// TIA Portal project "XSFW_TIA32801_A0" (V15.1)

(* hardware
DEVICE "Estación SIMATIC 1200_1"  S71200.Device
   slot 0: "Rack S7-1200"  Rack  V1.0
   slot 1: "PLC_1"  CPU 1214C DC/DC/DC  6ES7 214-1AG40-0XB0  V4.3
   slot 2: "DI16/DQ16 x 24V DC_1"  6ES7 223-1BL30-0XB0  V1.0
   slot 3: "DI 8x24VDC_1"  6ES7 221-1BF32-0XB0  V2.0
DEVICE "HMI_1"  KTP700 Basic PN
   slot 0: "HMI_1"  KTP700 Basic PN  6AV2 123-2GB03-0AX0  15.1.0.0
   slot 1: "HMI_RT_1"  KTP700 Basic PN  6AV2 123-2GB03-0AX0  15.1.0.0
   slot 5: "IE_CP_1"  PROFINET Interface  IE_CP  15.0.1.0
      slot 1: "PROFINET_Interfaz_1"  PROFINET Interface
         slot 1: "PORT_1"  Port  1.0.0.0
*)

// ===== PLC "PLC_1"  CPU 1214C DC/DC/DC =====

VAR_GLOBAL   // PLC tag table "Constantes del sistema"
   "Encoder" AT %ID1000 : DWord;   // Almacena el valor actual del encoder
   "System_Byte" AT %MB61 : Byte;
   "Clock_Byte" AT %MB60 : Byte;
   "Marca del sistema" AT %M61.0 : Bool;   // marca del sistema
   "Marca de ciclo" AT %M60.0 : Bool;   // Genera una luz titilante de 10 hz
   "No entrega caja" AT %M100.0 : Bool;
   "No libera salida" AT %M100.1 : Bool;
   "HMI_Hab. Falla caja trab." AT %M100.2 : Bool;
   "Tag_4" AT %M100.3 : Bool;
   "Tag_5" AT %M100.4 : Bool;
   "Tag_6" AT %M100.5 : Bool;
   "Tag_7" AT %M100.6 : Bool;
   "Tag_8" AT %M100.7 : Bool;
   "Tag_9" AT %M101.0 : Bool;
   "bit 1 de Reg_A" AT %M101.1 : Bool;
   "Tag_11" AT %M101.2 : Bool;
   "Tag_12" AT %M101.3 : Bool;
   "Tag_13" AT %M101.4 : Bool;
   "Tag_14" AT %M101.5 : Bool;
   "Tag_15" AT %M101.6 : Bool;
   "Tag_16" AT %M101.7 : Bool;
   "bit 0 de Reg_B" AT %M102.0 : Bool;
   "Tag_18" AT %M102.1 : Bool;
   "Tag_19" AT %M102.2 : Bool;
   "Tag_20" AT %M102.3 : Bool;
   "Tag_21" AT %M102.4 : Bool;
   "Tag_22" AT %M102.5 : Bool;
   "Tag_23" AT %M102.6 : Bool;
   "Tag_24" AT %M102.7 : Bool;
   "Tag_25" AT %M103.0 : Bool;
   "Tag_26" AT %M103.1 : Bool;
   "Tag_27" AT %M103.2 : Bool;
   "Tag_28" AT %QB0 : Byte;
   "UNO" AT %M27.0 : Bool;
   "CERO" AT %M27.1 : Bool;
   "Marca ciclo alim cartones" AT %M60.1 : Bool;   // es una marca de ciclo de 5 hz para manejar el alim de cartones
   "Tag_29" AT %M60.2 : Bool;
   "Tag_30" AT %M60.5 : Bool;
   "Tag_31" AT %MD300 : DWord;
   "Valor encoder pusher salida" AT %MD350 : DWord;
   "Tag_32" AT %E0.7 : Bool;
   "Tag_33" AT %M36.4 : Bool;
   "Reg_A" AT %MB101 : Byte;
   "Reg_B" AT %MB102 : Byte;
   "Tag_1" AT %I34.2 : Bool;
END_VAR

VAR_GLOBAL   // PLC tag table "Pusher"
   "iSNSpush_atras" AT %I33.2 : Bool;   // Detecta Pusher atrás
   "iSNSpush_adel" AT %I0.2 : Bool;   // Detecta Pusher adelante
   "iSNSalp" AT %I1.0 : Bool;   // Sensor área de recorrido libre del pusher
   "oM_pusher" AT %Q32.3 : Bool;   // Activa el pusher
   "oPusher_out" AT %Q33.5 : Bool;   // Activa válvula del Cilindro del pusher
END_VAR

VAR_GLOBAL   // PLC tag table "brazo de succion"
   "iSNS_bs_abajo" AT %I33.6 : Bool;   // Detecta cuando el brazo de succión está abajo
   "iSNS_bs_arriba" AT %I33.7 : Bool;   // Detecta cuando el brazo de succión está arriba
   "oM_brazo_succión" AT %Q32.2 : Bool;   // Activa el brazo de succión
   "oVálvula_Succión" AT %Q33.0 : Bool;   // Activa valvula chupetes succionadores
END_VAR

VAR_GLOBAL   // PLC tag table "Pinza"
   "oPinza" AT %Q33.6 : Bool;   // Activa válvula Brazos tipo pinza que cierran las solapas inferiores de la caja
END_VAR

VAR_GLOBAL   // PLC tag table "agarra solapa, cierra solapa, alimentador de caja,retenedores"
   "oAgarra_solapas" AT %Q33.1 : Bool;   // Activa válvula brazos agarra solapas
   "oCierra_solapa" AT %Q33.2 : Bool;   // Activa válvula brazo cierra solapa
   "oRetB" AT %Q33.3 : Bool;   // Activa válvula Retenedor de caja en sector B
   "oRetC" AT %Q33.7 : Bool;   // Activa válvula Retenedor de cajas en sector C
   "oAlim_cart" AT %Q0.0 : Bool;   // Válvula Alimentación automática de cartones
   "iSNS_nivel_bajo_cartones" AT %I33.0 : Bool;   // Detecta nivel bajo de cartones
END_VAR

VAR_GLOBAL   // PLC tag table "Encoladora"
   "iSNS_carton en area de colado" AT %I33.3 : Bool;   // Detecta el cartón en sector de colado
   "iK_encol_on" AT %I33.1 : Bool;   // Encoladora encendida y caliente (tarda 45 min en calentar)
   "iSNSpegamento en depósito" AT %I1.2 : Bool;   // Detecta pegamento en depósito
   "oBoquilla_Encoladora" AT %Q33.4 : Bool;   // Activa Boquilla encoladora
END_VAR

VAR_GLOBAL   // PLC tag table "Area de salida"
   "iSNScaja_trab" AT %I1.4 : Bool;   // Detecta cuando la caja cae a la cinta de salida
   "iSnsCajaCerrada" AT %I1.5 : Bool;   // Detecta si la caja no se abrio cuando bajo a la cadena
   "oM_cinta_sal" AT %Q32.4 : Bool;   // Activa la cinta de salida
   "iSNScaja_acum" AT %I0.4 : Bool;   // detecta cajas acumuladas
END_VAR

VAR_GLOBAL   // PLC tag table "Cinta y encoder"
   "iFaseA" AT %I0.0 : Bool;   // fase A del encoder
   "iFaseB" AT %I0.1 : Bool;   // fase B del encoder
   "iFase0" AT %I0.3 : Bool;   // fase 0 del encoder, detecta cuando se cumplió una vuelta
   "oM_cinta_principal" AT %Q32.0 : Bool;   // Activa el motor de la cinta principal
END_VAR

VAR_GLOBAL   // PLC tag table "auxiliares para almacenar flancos"
   "Guarda flanco subida caja acum" AT %M80.0 : Bool;   // almacena valor anterior del sensor caja acumulada
   "Guarda flanco bajada caja acum" AT %M80.1 : Bool;   // almacena valor anterior del sensor caja acumulada
   "Guarda flanco bajada caja trab" AT %M80.2 : Bool;   // almacena valor anterior del sensor caja trabada
   "Guarda flanco subida caja trab" AT %M80.3 : Bool;   // almacena valor anterior del sensor caja trabada
   "Guarda flanco brazo succión arriba" AT %M80.4 : Bool;   // Almacena el estado anterior del sensor
   "Guarda flanco subida area encolado" AT %M80.5 : Bool;
   "Guarda flanco bajada area encolado" AT %M80.6 : Bool;
   "Guarda flanco pulsador averia/reposicion" AT %M80.7 : Bool;
   "Guarda flanco subida pulsador marcha" AT %M81.0 : Bool;
   "Guarda flanco subida pulsador avería/reposición" AT %M81.1 : Bool;
   "Guarda flanco subida pulsador Parada" AT %M81.2 : Bool;
   "fls_Averiarep" AT %M81.3 : Bool;
   "fls_M" AT %M81.4 : Bool;
   "fls_Area_encol_sub" AT %M81.5 : Bool;
   "fls_Area_encol_baj" AT %M81.6 : Bool;
   "Guarda flanco Marcha desde panel" AT %M81.7 : Bool;
   "Guarda flanco modo manual" AT %M82.0 : Bool;
   "fls_Modomanual" AT %M82.1 : Bool;   // Pulsador desde panel para comenzar modo manual
   "Guarda flanco bajada alim cart" AT %M82.2 : Bool;
   "Guarda flanco de bajada sns brazo abajo" AT %M82.3 : Bool;
END_VAR

VAR_GLOBAL   // PLC tag table "Pulsadores y selectores"
   "iM" AT %I32.5 : Bool;   // Pulsador de Marcha
   "iP" AT %I32.6 : Bool;   // Pulsador de Parada
   "iS_automat" AT %I33.4 : Bool;   // Selector modo automático
   "iS_Probar" AT %I33.5 : Bool;   // Selector modo test
   "iS_cinta_salida_on" AT %I1.3 : Bool;   // Selectora on/off de la cinta de salida
END_VAR

VAR_GLOBAL   // PLC tag table "Seguridad"
   "iEmergencia" AT %I32.1 : Bool;   // Ventanas cerradas y emerg off
   "iAveria-reposicion" AT %I32.2 : Bool;   // Repone avería
   "iTermicas_mev" AT %I32.3 : Bool;   // Térmicas del motor, encoladora, bomba
   "iTermicas_pbs" AT %I32.4 : Bool;   // Térmicas del brazo de succión y pusher
   "iSNSproteccion_torque" AT %I0.5 : Bool;   // Sensor Protección de torque motor principal cinta
   "oLinea-emergencia" AT %Q32.7 : Bool;   // Salida a línea de emergencia
END_VAR

VAR_GLOBAL   // PLC tag table "voltage de control"
   "iEnable" AT %I32.0 : Bool;   // Voltage de control
END_VAR

VAR_GLOBAL   // PLC tag table "Otros"
   "k_EXT" AT %I1.1 : Bool;   // enable suction arm from EXT input
   "oQuick_out" AT %Q0.1 : Bool;   // ?
   "oSep_fing" AT %Q0.4 : Bool;   // ?
   "oPacker" AT %Q0.3 : Bool;   // En teoría se habilita luego que pulsa Marcha
   "desactivar" AT %M50.0 : Bool;
END_VAR

VAR_GLOBAL   // PLC tag table "Bomba de vacio"
   "oM_bomba" AT %Q32.1 : Bool;   // Activa la bomba de vacío
END_VAR

VAR_GLOBAL   // PLC tag table "Luces"
   "oLmpR" AT %Q32.5 : Bool;   // Lámpara para indicar parada y fallas de cualquier índole
   "oLmpV" AT %Q32.6 : Bool;   // Lámpara para indicar marcha
END_VAR

VAR_GLOBAL   // PLC tag table "Estados"
   "DS1" AT %MD0 : DWord;   // Variable tipo Word. Almacena los 12 Estados del proceso
   "1s1" AT %M0.0 : Bool;   // Estado 1: Reposo
   "1s2" AT %M0.1 : Bool;   // Estado 2: Activa Cinta ppal
   "1s3" AT %M0.2 : Bool;   // Estado 3: Activar retenedores de caja
   "1s4" AT %M0.3 : Bool;   // Estado 4: Desactivar Cinta ppal
   "1s5" AT %M0.4 : Bool;   // Estado 5: Activar Pusher y Pinza
   "1s6" AT %M0.5 : Bool;   // Estado 6: Activar Cilindro neumático Pusher
   "1s7" AT %M0.6 : Bool;   // Estado 7: Desactivar Pinza y Cilindro Pusher
   "1s8" AT %M0.7 : Bool;   // Estado 8: Área libre de Pusher
   "1s9" AT %M1.0 : Bool;   // Estado 9: Fin Etapa Pusher
   "1s10" AT %M1.1 : Bool;
   "1s11" AT %M1.2 : Bool;
   "1s12" AT %M1.3 : Bool;
   "DS2" AT %MD4 : DWord;
   "2s1" AT %M4.0 : Bool;   // Estado 8: Activar retenedores de caja
   "2s2" AT %M4.1 : Bool;   // Estado 9: Desactivar cinta
   "2s3" AT %M4.2 : Bool;   // Estado 10: Activa Pusher, Pinza y Cierra solapa
   "2s4" AT %M4.3 : Bool;   // Estado 11: Cilindro Pusher Afuera
   "2s5" AT %M4.4 : Bool;   // Estado 12: Desactivar Cilindro Pusher, Pinza y Cierra solapa
   "2s6" AT %M4.5 : Bool;   // Estado 13: Fin Pusher
   "2s7" AT %M4.6 : Bool;   // Estado 14: Area liberada del Pusher
   "2s8" AT %M4.7 : Bool;
   "2s9" AT %M5.0 : Bool;
   "2s10" AT %M5.1 : Bool;
   "2s11" AT %M5.2 : Bool;
   "2s12" AT %M5.3 : Bool;
   "2s13" AT %M5.4 : Bool;
   "2s14" AT %M5.5 : Bool;
   "2s15" AT %M5.6 : Bool;
   "2s16" AT %M5.7 : Bool;
   "2s17" AT %M6.0 : Bool;
   "2s18" AT %M6.1 : Bool;
   "2s19" AT %M6.2 : Bool;
   "2s20" AT %M6.3 : Bool;
   "2s21" AT %M6.4 : Bool;
   "2s22" AT %M6.5 : Bool;
   "2s23" AT %M6.6 : Bool;
   "2s24" AT %M6.7 : Bool;
   "2s25" AT %M7.0 : Bool;
   "2s26" AT %M7.1 : Bool;
   "2s27" AT %M7.2 : Bool;
   "2s28" AT %M7.3 : Bool;
   "2s29" AT %M7.4 : Bool;
   "2s30" AT %M7.5 : Bool;
   "2s31" AT %M7.6 : Bool;
   "2s32" AT %M7.7 : Bool;
   "1s13" AT %M1.4 : Bool;
   "1s14" AT %M1.5 : Bool;
   "1s15" AT %M1.6 : Bool;
   "1s16" AT %M1.7 : Bool;
   "1s17" AT %M2.0 : Bool;
   "1s18" AT %M2.1 : Bool;
   "1s19" AT %M2.2 : Bool;
   "1s20" AT %M2.3 : Bool;   // Estado de Alarmas
   "1s21" AT %M2.4 : Bool;   // Estado de parada
   "1s22" AT %M2.5 : Bool;   // Cajas acumuladas
   "1s23" AT %M2.6 : Bool;
   "1s24" AT %M2.7 : Bool;
   "1s25" AT %M3.0 : Bool;
   "1s26" AT %M3.1 : Bool;
   "1s27" AT %M3.2 : Bool;
   "1s28" AT %M3.3 : Bool;
   "1s29" AT %M3.4 : Bool;
   "1s30" AT %M3.5 : Bool;
   "1s31" AT %M3.6 : Bool;
   "1s32" AT %M3.7 : Bool;
END_VAR

VAR_GLOBAL   // PLC tag table "Concatenadores"
   "DC1" AT %MD8 : DWord;
   "1c1" AT %M8.0 : Bool;   // Ir a Estado 1: Reposo
   "1c2" AT %M8.1 : Bool;   // Ir a estado 2: Activa Cinta ppal
   "1c3" AT %M8.2 : Bool;   // Ir a estado 3: Activar retenedores de caja
   "1c4" AT %M8.3 : Bool;   // Ir estado 4: Desactivar Cinta ppal
   "1c5" AT %M8.4 : Bool;   // Ir a estado 5: Activar Pusher y Pinza
   "1c6" AT %M8.5 : Bool;   // Ir a estado 6: Activar cilindro neumático Pusher
   "1c7" AT %M8.6 : Bool;   // Ir a estado 7: Desactivar Pinza y Cilindro Pusher
   "DC2" AT %MD12 : DWord;
   "2c1" AT %M12.0 : Bool;   // Ir a Estado 8: Activar retenedores de caja
   "2c2" AT %M12.1 : Bool;   // Ir a Estado 9: Desactivar cinta
   "2c3" AT %M12.2 : Bool;   // Ir a Estado 10: Activa Pusher, Pinza y Cierra solapa
   "2c4" AT %M12.3 : Bool;   // Ir a Estado 11: Cilindro Pusher afuera
   "2c5" AT %M12.4 : Bool;   // Ir a Estado 12: Desactivar Cilindro Pusher, Pinza y Cierra solapa
   "2c6" AT %M12.5 : Bool;   // Ir a Estado 13: Fin Pusher
   "2c7" AT %M12.6 : Bool;   // Ir a Estado 14: Area liberada del Pusher
   "1c8" AT %M8.7 : Bool;   // Ir a Estado 8: Área libre de Pusher
   "1c9" AT %M9.0 : Bool;   // Ir a Estado 9: Fin etapa Pusher
   "1c10" AT %M9.1 : Bool;
   "1c11" AT %M9.2 : Bool;
   "1c12" AT %M9.3 : Bool;
   "1c13" AT %M9.4 : Bool;
   "1c14" AT %M9.5 : Bool;
   "1c15" AT %M9.6 : Bool;
   "1c16" AT %M9.7 : Bool;
   "1c17" AT %M10.0 : Bool;
   "1c18" AT %M10.1 : Bool;
   "1c19" AT %M10.2 : Bool;
   "1c20" AT %M10.3 : Bool;
   "1c21" AT %M10.4 : Bool;
   "1c22" AT %M10.5 : Bool;
   "1c23" AT %M10.6 : Bool;
   "1c24" AT %M10.7 : Bool;
   "1c25" AT %M11.0 : Bool;
   "1c26" AT %M11.1 : Bool;
   "1c27" AT %M11.2 : Bool;
   "1c28" AT %M11.3 : Bool;
   "1c29" AT %M11.4 : Bool;
   "1c30" AT %M11.5 : Bool;
   "1c31" AT %M11.6 : Bool;
   "1c32" AT %M11.7 : Bool;
   "2c8" AT %M12.7 : Bool;
   "2c9" AT %M13.0 : Bool;
   "2c10" AT %M13.1 : Bool;
   "2c11" AT %M13.2 : Bool;
   "2c12" AT %M13.3 : Bool;
   "2c13" AT %M13.4 : Bool;
   "2c14" AT %M13.5 : Bool;
   "2c15" AT %M13.6 : Bool;
   "2c16" AT %M13.7 : Bool;
   "2c17" AT %M14.0 : Bool;
   "2c18" AT %M14.1 : Bool;
   "2c19" AT %M14.2 : Bool;
   "2c20" AT %M14.3 : Bool;
   "2c21" AT %M14.4 : Bool;
   "2c22" AT %M14.5 : Bool;
   "2c23" AT %M14.6 : Bool;
   "2c24" AT %M14.7 : Bool;
   "2c25" AT %M15.0 : Bool;
   "2c26" AT %M15.1 : Bool;
   "2c27" AT %M15.2 : Bool;
   "2c28" AT %M15.3 : Bool;
   "2c29" AT %M15.4 : Bool;
   "2c30" AT %M15.5 : Bool;
   "2c31" AT %M15.6 : Bool;
   "2c32" AT %M15.7 : Bool;
END_VAR

VAR_GLOBAL   // PLC tag table "Marcas"
   "Marcha" AT %M20.0 : Bool;   // marca "Iniciar proceso"
   "Activar desplazador" AT %M20.1 : Bool;   // marca "activar cilindro alimentador"
   "Activa_cinta_salida" AT %M20.2 : Bool;   // marca " activa cinta de salida"
   "HMI_Hab_Falla_Caja_Caida" AT %M20.3 : Bool;   // Cajas acumuladas en la cinta de salida
   "Interrumpir" AT %M20.4 : Bool;   // Interrumpe el proceso
   "Activa pinza" AT %M20.5 : Bool;   // Activa la pinza
   "Activa cierra solapa" AT %M20.6 : Bool;   // Activa el cierra solapa
   "Activa bomba" AT %M20.7 : Bool;   // Activa la bomba de vacío
   "Activa brazo_succion" AT %M21.0 : Bool;   // Activa el motor del brazo de succión
   "Pusher-atras-ok" AT %M21.2 : Bool;   // Confirma que el pusher tocó el sensor de atrás
   "Pusher-adelante-ok" AT %M21.3 : Bool;   // Confirma que el pusher tocó el sensor adelante
   "Area libre del pusher" AT %M21.4 : Bool;   // Confirma que se activó el sensor
   "Ya buscó caja" AT %M21.5 : Bool;   // Confirma que el brazo tomó una caja
   "Activa succionadores" AT %M21.6 : Bool;   // Marca que activa los chupetes succionadores
   "No salió caja" AT %M21.7 : Bool;   // Indica que la caja no salió del rango del brazo de succión
   "Aux1" AT %M22.0 : Bool;   // auxiliar para los registros SR
   "Aux2" AT %M22.1 : Bool;   // auxiliar para los registros SR
   "Aux3" AT %M22.2 : Bool;   // auxiliar para los registros SR
   "Aux4" AT %M22.3 : Bool;   // auxiliar para los registros SR
   "Aux5" AT %M22.4 : Bool;   // auxiliar para los registros SR
   "Encolado fallido o falla en sensor" AT %M23.0 : Bool;   // Indica que el encolado se realizó correctamente, se da cuuando NO se da falla en encolado
   "Rearmar" AT %M23.1 : Bool;   // Se activa cuando se presiona el pulsador de avería/reposición
   "Falla en pusher" AT %M23.2 : Bool;   // Indica que hubo una falla en el pusher
   "Alarmas pusher" AT %M23.3 : Bool;   // Agrupa las alarmas del pusher
   "Alarmas brazo de succión" AT %M23.4 : Bool;   // Agrupa las alarmas del brazo de succión
   "Alarmas emergencia y térmicas" AT %M23.5 : Bool;   // Agrupa las alarmas de la serie térmicas y serie emergencia y ventanas
   "Alarmas cinta" AT %M23.6 : Bool;   // Agrupa las alarmas de la cinta
   "Alarmas salida y alim de cartones" AT %M23.7 : Bool;   // Agrupa las alarmas de la salida de la máquina (caja trabada) y alimentación de cartones
   "Cajas acumuladas en salida" AT %M24.0 : Bool;   // Detecta acumulación de cajas en la cinta salida interrumpiendo el proceso
   "Aux6" AT %M24.1 : Bool;
   "Alarmas encoladora" AT %M24.2 : Bool;
   "Serie de Alarmas" AT %M24.3 : Bool;
   "Habilita modo Probar" AT %M24.4 : Bool;
   "Tiempo de encolado solapa 1" AT %M24.5 : Bool;
   "Tiempo de encolado solapa2" AT %M24.6 : Bool;
   "Serie de fallas" AT %M24.7 : Bool;
   "Rearme desde panel" AT %M25.0 : Bool;
   "Emergencia desde panel" AT %M25.1 : Bool;
   "Valor del encoder" AT %MD180 : DWord;
   "Parada" AT %M25.2 : Bool;
   "Marcha desde panel" AT %M25.3 : Bool;
   "Modo Manual" AT %M25.4 : Bool;   // Cuando no está en modo probar ni en modo aut, está en modo manual
   "Resetear cajas armadas" AT %M25.5 : Bool;
   "Valor cantidad de cajas armadas" AT %MD120 : DWord;
   "Valor de referencia cajas armadas" AT %M25.6 : Bool;
   "Aux7" AT %M25.7 : Bool;
   "Solapa en área de encolado" AT %M26.0 : Bool;
   "Solapa fuera del area de encolado" AT %M26.1 : Bool;
   "Valorexp de contaje para calcular encolado x" AT %MD150 : DWord;
   "Exp Almacena el valor encolado experimental" AT %MD170 : DWord;
   "Exp marca de prueba fase 0" AT %M26.2 : Bool;   // Esta marca sólo me sirve a mi para ver si la fase 0 efectiv se activa
   "Impedir falla" AT %M26.3 : Bool;
   "Boton activar fingers" AT %M26.4 : Bool;
   "Botón packer" AT %M26.5 : Bool;
   "Boton quick out" AT %M26.6 : Bool;
   "Exp valor del encoder para calc encolado" AT %MD220 : DWord;
   "Exp marca aux id118" AT %M22.5 : Bool;
   "Pulsador modo manual" AT %M22.6 : Bool;   // Cada vez que se pulsa, se lleva a cabo un ciclo de la armadora
   "Aviso de cinta descalibrada probar" AT %M22.7 : Bool;
   "Habilitar brazo manual" AT %M26.7 : Bool;
   "Aux alim cart" AT %M27.2 : Bool;
   "Aux alim cart 2" AT %M27.3 : Bool;
   "Iniciar temp alim cart" AT %M27.4 : Bool;
   "Recuerda paso pusher" AT %M27.5 : Bool;
   "Auxiliar encoder exp" AT %M27.6 : Bool;
   "Aux9" AT %M27.7 : Bool;
   "Punto neutro" AT %M28.0 : Bool;
   "Aux10" AT %M28.1 : Bool;
   "Aux11" AT %M28.2 : Bool;
   "Delay cierra solapa" AT %M28.3 : Bool;
   "Delay brazo" AT %M28.4 : Bool;
   "Delay brazo 2" AT %M28.5 : Bool;
   "Aux12" AT %M28.6 : Bool;
   "Auxencol1" AT %M28.7 : Bool;
   "Auxencol2" AT %M29.0 : Bool;
   "Guarda flanco bajada averi rep delay" AT %M29.1 : Bool;
   "Rearme delay" AT %M29.2 : Bool;
   "Delaymarcha" AT %M29.3 : Bool;
   "Guarda flanco delay  marcha" AT %M29.4 : Bool;
   "Parar proceso" AT %M29.5 : Bool;
   "Espera caja" AT %M29.6 : Bool;
   "Guarda flanco punto m" AT %M29.7 : Bool;
   "Parar brazo" AT %M34.0 : Bool;
   "Flanco 2" AT %M34.1 : Bool;
   "Esperar cinta" AT %M34.2 : Bool;
   "Flanco p atras" AT %M34.3 : Bool;
   "Flanco nivel bajo" AT %M34.4 : Bool;
   "Retrasa nivel bajo c" AT %M34.5 : Bool;
   "Fls sns b abajo" AT %M34.6 : Bool;
   "Fls_bajada snsalp" AT %M34.7 : Bool;
   "Aux marca pusher" AT %M35.0 : Bool;
   "Aux acaja acum" AT %M35.1 : Bool;
   "Aux17" AT %M35.2 : Bool;
   "Aux caja trab" AT %M35.3 : Bool;
   "Marca aux" AT %M35.4 : Bool;
   "Fsnsalp" AT %M35.5 : Bool;
   "Xsnsalp" AT %M35.6 : Bool;
   "FallaSnsAtras" AT %M35.7 : Bool;
   "F1s8" AT %M36.0 : Bool;
   "X1s8" AT %M36.1 : Bool;
   "Flanco_PusherAtras" AT %M36.2 : Bool;
   "FlancoAtras_Detectado" AT %M36.3 : Bool;
END_VAR

VAR_GLOBAL   // PLC tag table "Prioritarias"
   "1p1" AT %M16.0 : Bool;
   "DP1" AT %MD16 : DWord;
   "1p2" AT %M16.1 : Bool;
   "1p3" AT %M16.2 : Bool;
   "1p4" AT %M16.3 : Bool;
   "DP2" AT %MD30 : DWord;
   "2p1" AT %M30.0 : Bool;
   "2p2" AT %M30.1 : Bool;
   "2p3" AT %M30.2 : Bool;
   "2p4" AT %M30.3 : Bool;
   "2p5" AT %M30.4 : Bool;
   "2p6" AT %M30.5 : Bool;
   "1p8" AT %M16.7 : Bool;
   "1p9" AT %M17.0 : Bool;
   "1p5" AT %M16.4 : Bool;
   "1p6" AT %M16.5 : Bool;
   "1p7" AT %M16.6 : Bool;
   "1p10" AT %M17.1 : Bool;
   "1p11" AT %M17.2 : Bool;
   "1p12" AT %M17.3 : Bool;
   "1p13" AT %M17.4 : Bool;
   "1p14" AT %M17.5 : Bool;
   "1p15" AT %M17.6 : Bool;
   "1p16" AT %M17.7 : Bool;
   "1p17" AT %M18.0 : Bool;
   "1p18" AT %M18.1 : Bool;
   "1p19" AT %M18.2 : Bool;
   "1p20" AT %M18.3 : Bool;   // Prioritaria que para el proceso y necesita rearme
   "1p21" AT %M18.4 : Bool;   // Prioritaria que para el proceso y no necesita rearme
   "1p22" AT %M18.5 : Bool;   // Cajas acumuladas
   "1p23" AT %M18.6 : Bool;
   "1p24" AT %M18.7 : Bool;
   "1p25" AT %M19.0 : Bool;
   "1p26" AT %M19.1 : Bool;
   "1p27" AT %M19.2 : Bool;
   "1p28" AT %M19.3 : Bool;
   "1p29" AT %M19.4 : Bool;
   "1p30" AT %M19.5 : Bool;
   "1p31" AT %M19.6 : Bool;
   "1p32" AT %M19.7 : Bool;
END_VAR

VAR_GLOBAL   // PLC tag table "Modo probar"
   "MPbrazo de succión arriba" AT %M40.0 : Bool;   // levanta el brazo de succión
   "MPbrazo de succión abajo" AT %M40.1 : Bool;
   "MPlevanta brazo" AT %M40.2 : Bool;
   "MPbaja brazo" AT %M40.3 : Bool;
   "MPbotón Activa succión" AT %M40.4 : Bool;
   "MPsucciona caja" AT %M40.6 : Bool;
   "MPboton Activar bomba de vacío" AT %M40.7 : Bool;
   "MPbotón Activar encoladora" AT %M41.0 : Bool;
   "MPtiempo de encolado" AT %M41.1 : Bool;   // Encola por 2 segundos, independientemente si sigo presionando el botón
   "MPbotón alimentador de cartones" AT %M41.2 : Bool;
   "MPbotón Agarra solapas" AT %M41.3 : Bool;
   "MPbotón Cierra solapa" AT %M41.4 : Bool;
   "MPbotón Avanzar cinta" AT %M41.5 : Bool;
   "MPvalor actual del encoder" AT %MD200 : DWord;
   "MPbotón Avanzar cinta por tramos" AT %M41.6 : Bool;
   "MPActivar cinta" AT %M41.7 : Bool;
   "MPbotón activar pusher" AT %M42.0 : Bool;
   "MPActivar pusher" AT %M42.1 : Bool;
   "MPActivar cilindro pusher" AT %M42.2 : Bool;
   "MPguarda flanco subida ALP" AT %M42.3 : Bool;
   "MPActivar pinza" AT %M42.4 : Bool;
   "MPActiva bomba de vacío" AT %M42.5 : Bool;
   "MPActiva encola" AT %M42.6 : Bool;
   "MPActiva alimentación cartones" AT %M42.7 : Bool;
   "MPActiva los agarra solapas" AT %M43.0 : Bool;
   "MPActiva el cierra solapa" AT %M43.1 : Bool;
   "MPActiva la cinta de salida de cajas" AT %M43.2 : Bool;
   "ModoProbar" AT %M43.3 : Bool;
   "MPbotón activar retenedores de caja" AT %M43.4 : Bool;
   "MPActiva retenedores de caja" AT %M43.5 : Bool;
   "MPAcomodar brazo de succión" AT %M43.6 : Bool;
   "MPReset cuenta modo probar" AT %M43.7 : Bool;
   "MPboton cilindro push" AT %M44.0 : Bool;
   "MPactivar cilindro push" AT %M44.1 : Bool;
END_VAR

DATA_BLOCK "Fallas"   // DB1
{ S7_Optimized_Access := 'FALSE' }
VERSION : 0.1
   VAR
      termicas1 : Bool;   // Térmicas de la bomba de vacío, motor ppal, encoladora.
      termicas2 : Bool;   // Térmicas brazo de succión y pusher.
      emergencia : Bool;   // Ventanas abiertas o pulsador de emergencia activado.
      "proteccion de torque" : Bool;   // Protección de torque motor ppal (atasco).
      "Falla en rele cadena" : Bool;   // Falla en sensor de caja en área de encolado.
      "Falla en sensores del Pusher" : Bool;   // Falla en sensor del pusher atrás
      "Sensor pusher hacia adelante" : Bool;   // Falla en sensor del pusher adelante
      falla_sns_bsucc_ar : Bool;   // Falla en sensor del brazo de succión arriba
      falla_sns_bsucc_ab : Bool;   // Falla en sensor del brazo de succión abajo
      "area de recorrido libre del pusher" : Bool;   // Falla en sensor del pusher área libre.
      falla_alim_cartones : Bool;   // Falla en sensor alimentador de cartones.
      falla_encoder : Bool;   // Falla en encoder
      "caja trabada a la salida" : Bool;   // Falla en sensor de caja trabada a la salida.
      "Incrongruencia pusher" : Bool;   // Incongruencia en sensores del pusher
      "Falla de programación prioritarias 1" : Bool;
      "Falla de programación concatenadoras 1" : Bool;
      "Falla de programación prioritarias 2" : Bool;
      "Falla de programación concatenadoras 2" : Bool;
      "Falla en sensor de encolado" : Bool;   // Falla en sensor área de encolado
      "Sin pegamento en el depósito" : Bool;   // Sin pegamento en el depósito
      "falla rele cadena" : Bool;
      "Falla de caja cerrada en cadena" : Bool;   // se activa si cae mal la caja
      "Reserva 1_2_1" : Bool;
      "Reserva 1_3_1" : Bool;
      "Reserva 1_4_1" : Bool;
      "Reserva 1_4_1_1" : Bool;
      "Reserva 1_4_1_2" : Bool;
      "Reserva 1_4_1_3" : Bool;
      "Reserva 1_4_1_4" : Bool;
      "Reserva 1_4_1_4_1" : Bool;
      "Reserva 1_4_1_4_1_1" : Bool;
      "Reserva 1_4_1_4_1_2" : Bool;
   END_VAR
BEGIN
END_DATA_BLOCK

DATA_BLOCK "HSC"   // DB4
{ S7_Optimized_Access := 'FALSE' }
VERSION : 0.1
   VAR
      "punto muerto" : Bool;   // Indica que la cinta está completamente detenida
      id118 : Bool;   // Cuando el encoder llega a contar 118 pulsos, apaga el motor
      "Se cumplio una vuelta" : Bool;   // Indica que el motor dió una vuelta completa
   END_VAR
BEGIN
END_DATA_BLOCK

DATA_BLOCK "datos de encolado"   // DB11
{ S7_Optimized_Access := 'FALSE' }
VERSION : 0.1
   VAR
      Iniciosol1cj1000 : DInt;
      finsol1cj1000 : DInt;
      Iniciosol2cj1000 : DInt;
      finsol2cj1000 : DInt;
      Iniciosol1cj1500 : DInt;
      finsol1cj1500 : DInt;
      Iniciosol2cj1500 : DInt;
      finsol2cj1500 : DInt;
      "selcaja1000/1500" : Bool;
   END_VAR
BEGIN
END_DATA_BLOCK

DATA_BLOCK "AjusteEncoder"   // DB17
{ S7_Optimized_Access := 'TRUE' }
VERSION : 0.1
   VAR
      Hab_Pusher : DInt := -10;   // 0
      Dhab_Pusher : DInt := 21;   // 21
      Reset_Val : DInt;
      Reset : Bool;
   END_VAR
BEGIN
END_DATA_BLOCK

DATA_BLOCK "Alarmas"   // DB19
{ S7_Optimized_Access := 'FALSE' }
VERSION : 0.1
   VAR
      termicas1 : Bool;   // Térmicas de la bomba de vacío, motor ppal, encoladora.
      termicas2 : Bool;   // Térmicas brazo de succión y pusher.
      emergencia : Bool;   // Ventanas abiertas o pulsador de emergencia activado.
      "proteccion de torque" : Bool;   // Protección de torque motor ppal (atasco).
      "falla en rele de cadena" : Bool;   // Falla en sensor de caja en área de encolado.
      "Falla en sensor atras del pusher" : Bool;   // Falla en sensor del pusher atrás
      "Sensor pusher hacia adelante" : Bool;   // Falla en sensor del pusher adelante
      falla_sns_bsucc_ar : Bool;   // Falla en sensor del brazo de succión arriba
      falla_sns_bsucc_ab : Bool;   // Falla en sensor del brazo de succión abajo
      "area de recorrido libre del pusher" : Bool;   // Falla en sensor del pusher área libre.
      falla_alim_cartones : Bool;   // Falla en sensor alimentador de cartones.
      falla_encoder : Bool;   // Falla en encoder
      "caja trabada a la salida" : Bool;   // Falla en sensor de caja trabada a la salida.
      "Incrongruencia pusher" : Bool;   // Incongruencia en sensores del pusher
      "Falla de programación prioritarias" : Bool;
      "Falla de programación concatenadoras" : Bool;
      "Falla de programación prioritarias 2" : Bool;
      "Falla de programación concatenadoras 2" : Bool;
      "Falla en sensor de encolado" : Bool;   // Falla en sensor área de encolado
      "Sin pegamento en el depósito" : Bool;   // Sin pegamento en el depósito
      "falla rele cadena" : Bool;
      "caja cerrada en cadena" : Bool;
      Reserva_9 : Bool;
      Reserva_10 : Bool;
      Reserva_11 : Bool;
      Reserva_12 : Bool;
      Reserva_13 : Bool;
      Reserva_14 : Bool;
      Reserva_15 : Bool;
      Reserva_15_1 : Bool;
      Reserva_15_1_1 : Bool;
      Reserva_15_1_2 : Bool;
   END_VAR
BEGIN
END_DATA_BLOCK

DATA_BLOCK "Tiempos"   // DB23
{ S7_Optimized_Access := 'FALSE' }
VERSION : 0.1
   VAR
      "Tiempo cierra sol" : DInt;
      "Tiempo espera brazo" : DInt;
      "tiempo cajas acum" : DInt;
      "Tiempo caja trabada" : DInt;
   END_VAR
BEGIN
END_DATA_BLOCK

// folder: System blocks/Program resources

DATA_BLOCK "Timer_DB2"   // DB2
{ S7_Optimized_Access := 'TRUE' }
AUTHOR : Simatic
FAMILY : IEC
NAME : IEC_TMR
VERSION : 1.0
// stored: InstanceOfName IEC_TIMER
"IEC_TIMER"
BEGIN
END_DATA_BLOCK

DATA_BLOCK "Timer_DB3"   // DB3
{ S7_Optimized_Access := 'TRUE' }
AUTHOR : Simatic
FAMILY : IEC
NAME : IEC_TMR
VERSION : 1.0
// stored: InstanceOfName IEC_TIMER
"IEC_TIMER"
BEGIN
END_DATA_BLOCK

DATA_BLOCK "Timer_DB5"   // DB5
{ S7_Optimized_Access := 'TRUE' }
AUTHOR : Simatic
FAMILY : IEC
NAME : IEC_TMR
VERSION : 1.0
// stored: InstanceOfName IEC_TIMER
"IEC_TIMER"
BEGIN
END_DATA_BLOCK

DATA_BLOCK "Timer_DB6"   // DB6
{ S7_Optimized_Access := 'TRUE' }
AUTHOR : Simatic
FAMILY : IEC
NAME : IEC_TMR
VERSION : 1.0
// stored: InstanceOfName IEC_TIMER
"IEC_TIMER"
BEGIN
END_DATA_BLOCK

DATA_BLOCK "Timer_DB7"   // DB7
{ S7_Optimized_Access := 'TRUE' }
AUTHOR : Simatic
FAMILY : IEC
NAME : IEC_TMR
VERSION : 1.0
// stored: InstanceOfName IEC_TIMER
"IEC_TIMER"
BEGIN
END_DATA_BLOCK

DATA_BLOCK "Timer_DB8"   // DB8
{ S7_Optimized_Access := 'TRUE' }
AUTHOR : Simatic
FAMILY : IEC
NAME : IEC_TMR
VERSION : 1.0
// stored: InstanceOfName IEC_TIMER
"IEC_TIMER"
BEGIN
END_DATA_BLOCK

DATA_BLOCK "Timer_DB9"   // DB9
{ S7_Optimized_Access := 'TRUE' }
AUTHOR : Simatic
FAMILY : IEC
NAME : IEC_TMR
VERSION : 1.0
// stored: InstanceOfName IEC_TIMER
"IEC_TIMER"
BEGIN
END_DATA_BLOCK

DATA_BLOCK "IEC_Timer_0_DB"   // DB10
{ S7_Optimized_Access := 'TRUE' }
AUTHOR : Simatic
FAMILY : IEC
NAME : IEC_TMR
VERSION : 1.0
// stored: InstanceOfName IEC_TIMER
"IEC_TIMER"
BEGIN
END_DATA_BLOCK

DATA_BLOCK "Timer_DB12"   // DB12
{ S7_Optimized_Access := 'TRUE' }
AUTHOR : Simatic
FAMILY : IEC
NAME : IEC_TMR
VERSION : 1.0
// stored: InstanceOfName IEC_TIMER
"IEC_TIMER"
BEGIN
END_DATA_BLOCK

DATA_BLOCK "Timer_DB13"   // DB13
{ S7_Optimized_Access := 'TRUE' }
AUTHOR : Simatic
FAMILY : IEC
NAME : IEC_TMR
VERSION : 1.0
// stored: InstanceOfName IEC_TIMER
"IEC_TIMER"
BEGIN
END_DATA_BLOCK

DATA_BLOCK "Timer_DB14"   // DB14
{ S7_Optimized_Access := 'TRUE' }
AUTHOR : Simatic
FAMILY : IEC
NAME : IEC_TMR
VERSION : 1.0
// stored: InstanceOfName IEC_TIMER
"IEC_TIMER"
BEGIN
END_DATA_BLOCK

DATA_BLOCK "Timer_DB15"   // DB15
{ S7_Optimized_Access := 'TRUE' }
AUTHOR : Simatic
FAMILY : IEC
NAME : IEC_TMR
VERSION : 1.0
// stored: InstanceOfName IEC_TIMER
"IEC_TIMER"
BEGIN
END_DATA_BLOCK

DATA_BLOCK "Contador_0"   // DB16
{ S7_Optimized_Access := 'TRUE' }
AUTHOR : SIMATIC
FAMILY : IEC
NAME : DCNTR
VERSION : 1.2
// stored: InstanceOfName IEC_DCOUNTER
"IEC_DCOUNTER"
BEGIN
END_DATA_BLOCK

DATA_BLOCK "Timer_DB18"   // DB18
{ S7_Optimized_Access := 'TRUE' }
AUTHOR : Simatic
FAMILY : IEC
NAME : IEC_TMR
VERSION : 1.0
// stored: InstanceOfName IEC_TIMER
"IEC_TIMER"
BEGIN
END_DATA_BLOCK

DATA_BLOCK "Timer_DB20"   // DB20
{ S7_Optimized_Access := 'TRUE' }
AUTHOR : Simatic
FAMILY : IEC
NAME : IEC_TMR
VERSION : 1.0
// stored: InstanceOfName IEC_TIMER
"IEC_TIMER"
BEGIN
END_DATA_BLOCK

DATA_BLOCK "Timer_DB21"   // DB21
{ S7_Optimized_Access := 'TRUE' }
AUTHOR : Simatic
FAMILY : IEC
NAME : IEC_TMR
VERSION : 1.0
// stored: InstanceOfName IEC_TIMER
"IEC_TIMER"
BEGIN
END_DATA_BLOCK

DATA_BLOCK "Timer_DB22"   // DB22
{ S7_Optimized_Access := 'TRUE' }
AUTHOR : Simatic
FAMILY : IEC
NAME : IEC_TMR
VERSION : 1.0
// stored: InstanceOfName IEC_TIMER
"IEC_TIMER"
BEGIN
END_DATA_BLOCK

DATA_BLOCK "Timer_DB24"   // DB24
{ S7_Optimized_Access := 'TRUE' }
AUTHOR : Simatic
FAMILY : IEC
NAME : IEC_TMR
VERSION : 1.0
// stored: InstanceOfName IEC_TIMER
"IEC_TIMER"
BEGIN
END_DATA_BLOCK

DATA_BLOCK "TOFF"   // DB26
{ S7_Optimized_Access := 'TRUE' }
AUTHOR : Simatic
FAMILY : IEC
NAME : IEC_TMR
VERSION : 1.0
// stored: InstanceOfName IEC_TIMER
"IEC_TIMER"
BEGIN
END_DATA_BLOCK

DATA_BLOCK "Desactivar Pusher"   // DB27
{ S7_Optimized_Access := 'TRUE' }
AUTHOR : Simatic
FAMILY : IEC
NAME : IEC_TMR
VERSION : 1.0
// stored: InstanceOfName IEC_TIMER
"IEC_TIMER"
BEGIN
END_DATA_BLOCK

DATA_BLOCK "Timer_DB30"   // DB30
{ S7_Optimized_Access := 'TRUE' }
AUTHOR : Simatic
FAMILY : IEC
NAME : IEC_TMR
VERSION : 1.0
// stored: InstanceOfName IEC_TIMER
"IEC_TIMER"
BEGIN
END_DATA_BLOCK

DATA_BLOCK "Timer_DB31"   // DB31
{ S7_Optimized_Access := 'TRUE' }
AUTHOR : Simatic
FAMILY : IEC
NAME : IEC_TMR
VERSION : 1.0
// stored: InstanceOfName IEC_TIMER
"IEC_TIMER"
BEGIN
END_DATA_BLOCK

// folder: (top level)

FUNCTION "Alimentador de cartones y cinta de salida" : Void   // FC1, LAD
TITLE = Desplaza una cinta que traslada los cartones hasta el brazo succionador.
{ S7_Optimized_Access := 'FALSE' }
VERSION : 0.1
BEGIN

REGION Network 1: Activa la cinta de salida
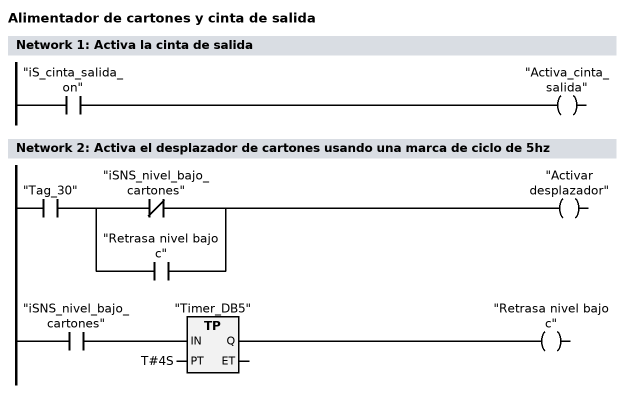
   RUNG wire#powerrail
      Contact( "iS_cinta_salida_on" )
      Coil( "Activa_cinta_salida" )
   END_RUNG
   // the same network as SCL:
   "Activa_cinta_salida" := "iS_cinta_salida_on";
END_REGION

REGION Network 2: Activa el desplazador de cartones usando una marca de ciclo de 5hz
   "Activar desplazador" := "Tag_30" AND (NOT "iSNS_nivel_bajo_cartones" OR "Retrasa nivel bajo c");
   "Timer_DB5".TP(IN := "iSNS_nivel_bajo_cartones", PT := T#4S);
   "Retrasa nivel bajo c" := "Timer_DB5".Q;
END_REGION
END_FUNCTION

FUNCTION "Tratamiento de Alarmas" : Void   // FC3, LAD
{ S7_Optimized_Access := 'TRUE' }
VERSION : 0.1
// Cada vez que ocurre una falla, cualquiera que fuese, se copia el estado de los bits de la doble palabra de "Fallas" a la doble palabra "Alarmas". Una vez resuelta la falla, se debe presionar "avería/reposición", lo cual generará un " reconocimiento de falla, que dará de baja la Alarma. A partir del segmento 4, agrupo las alarmas por función. Un grupo de alarmas para el pusher, uno para brazo de succión ,etc.
   VAR_TEMP
      "Alarmas presentes" : Word;
      Reconocimiento : Word;
   END_VAR
BEGIN

REGION Network 1: Reconocimiento/Reposición
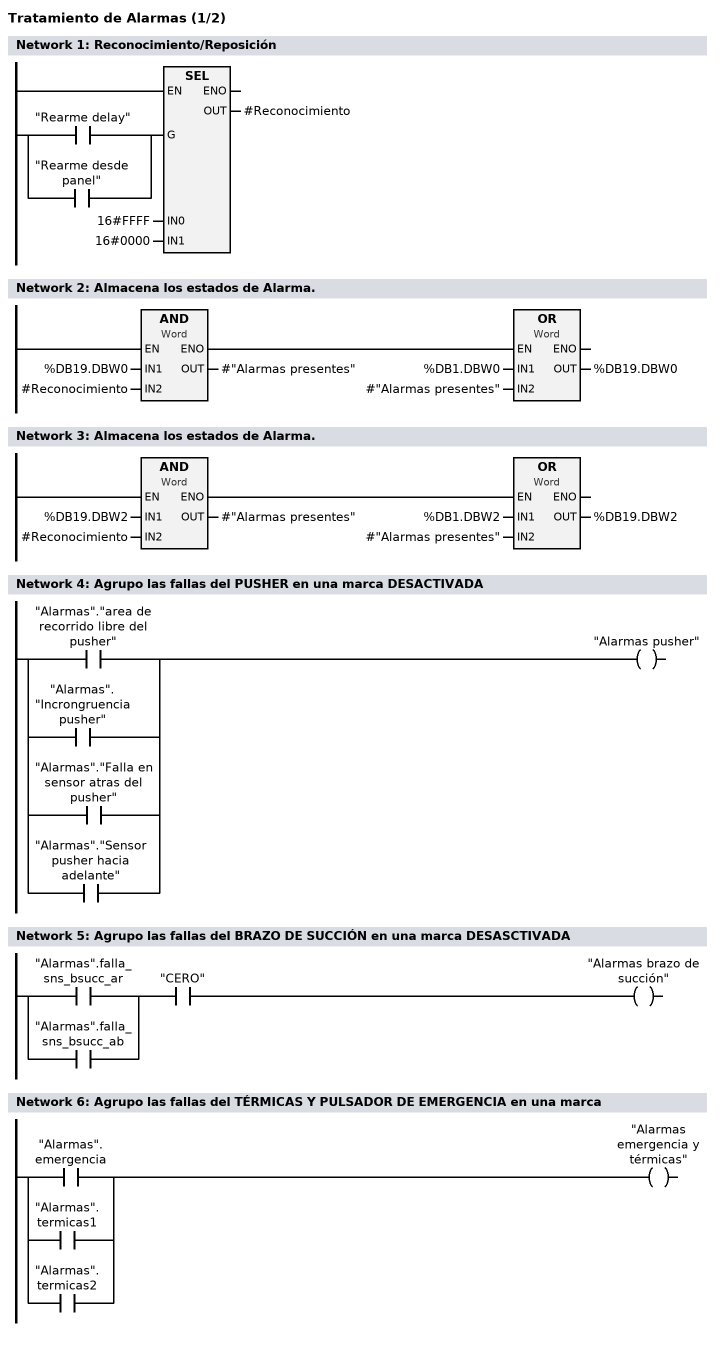
   #Reconocimiento := SEL(G := "Rearme delay" OR "Rearme desde panel", IN0 := 16#FFFF, IN1 := 16#0000);
END_REGION

REGION Network 2: Almacena los estados de Alarma.
   #"Alarmas presentes" := %DB19.DBW0 AND #Reconocimiento;
   %DB19.DBW0 := %DB1.DBW0 OR #"Alarmas presentes";
END_REGION

REGION Network 3: Almacena los estados de Alarma.
   #"Alarmas presentes" := %DB19.DBW2 AND #Reconocimiento;
   %DB19.DBW2 := %DB1.DBW2 OR #"Alarmas presentes";
END_REGION

REGION Network 4: Agrupo las fallas del PUSHER en una marca DESACTIVADA
   RUNG wire#powerrail
      Contact( "Alarmas"."area de recorrido libre del pusher" )
      wire#w1
      Coil( "Alarmas pusher" )
   END_RUNG
   RUNG wire#powerrail
      Contact( "Alarmas"."Incrongruencia pusher" )
   END_RUNG wire#w1
   RUNG wire#powerrail
      Contact( "Alarmas"."Falla en sensor atras del pusher" )
   END_RUNG wire#w1
   RUNG wire#powerrail
      Contact( "Alarmas"."Sensor pusher hacia adelante" )
   END_RUNG wire#w1
   // the same network as SCL:
   "Alarmas pusher" := "Alarmas"."area de recorrido libre del pusher" OR "Alarmas"."Incrongruencia pusher" OR "Alarmas"."Falla en sensor atras del pusher" OR "Alarmas"."Sensor pusher hacia adelante";
END_REGION

REGION Network 5: Agrupo las fallas del BRAZO DE SUCCIÓN en una marca DESASCTIVADA
   RUNG wire#powerrail
      Contact( "Alarmas".falla_sns_bsucc_ar )
      wire#w1
      Contact( "CERO" )
      Coil( "Alarmas brazo de succión" )
   END_RUNG
   RUNG wire#powerrail
      Contact( "Alarmas".falla_sns_bsucc_ab )
   END_RUNG wire#w1
   // the same network as SCL:
   "Alarmas brazo de succión" := ("Alarmas".falla_sns_bsucc_ar OR "Alarmas".falla_sns_bsucc_ab) AND "CERO";
END_REGION

REGION Network 6: Agrupo las fallas del TÉRMICAS Y PULSADOR DE EMERGENCIA en una marca
   RUNG wire#powerrail
      Contact( "Alarmas".emergencia )
      wire#w1
      Coil( "Alarmas emergencia y térmicas" )
   END_RUNG
   RUNG wire#powerrail
      Contact( "Alarmas".termicas1 )
   END_RUNG wire#w1
   RUNG wire#powerrail
      Contact( "Alarmas".termicas2 )
   END_RUNG wire#w1
   // the same network as SCL:
   "Alarmas emergencia y térmicas" := "Alarmas".emergencia OR "Alarmas".termicas1 OR "Alarmas".termicas2;
END_REGION

REGION Network 7: Agrupo las fallas de la CINTA en una marca
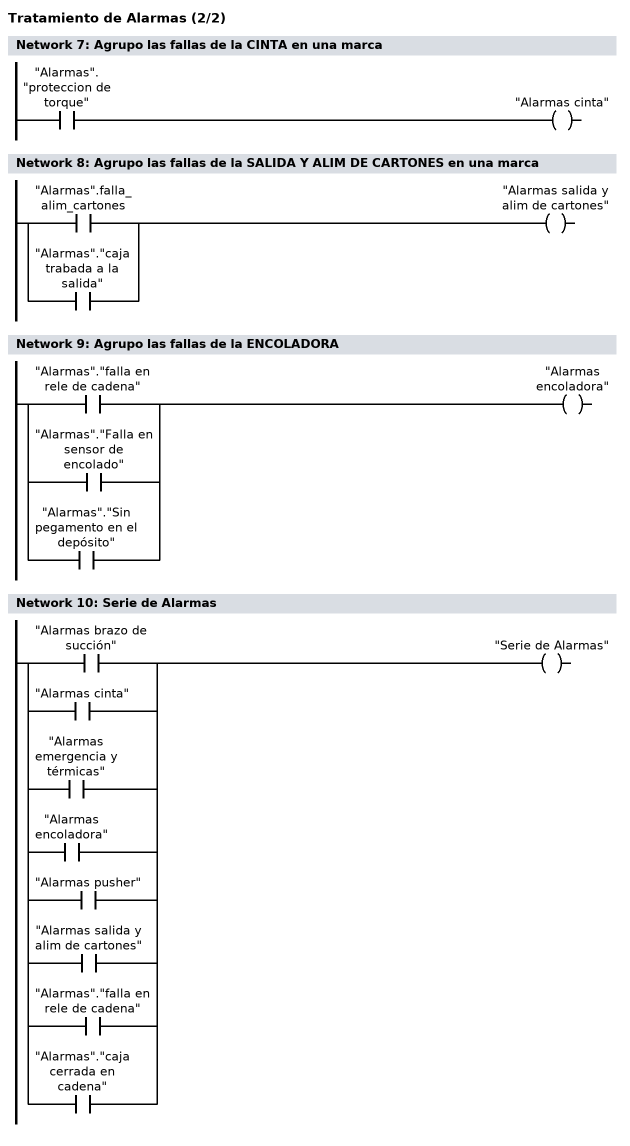
   RUNG wire#powerrail
      Contact( "Alarmas"."proteccion de torque" )
      Coil( "Alarmas cinta" )
   END_RUNG
   // the same network as SCL:
   "Alarmas cinta" := "Alarmas"."proteccion de torque";
END_REGION

REGION Network 8: Agrupo las fallas de la SALIDA Y ALIM DE CARTONES en una marca
   RUNG wire#powerrail
      Contact( "Alarmas".falla_alim_cartones )
      wire#w1
      Coil( "Alarmas salida y alim de cartones" )
   END_RUNG
   RUNG wire#powerrail
      Contact( "Alarmas"."caja trabada a la salida" )
   END_RUNG wire#w1
   // the same network as SCL:
   "Alarmas salida y alim de cartones" := "Alarmas".falla_alim_cartones OR "Alarmas"."caja trabada a la salida";
END_REGION

REGION Network 9: Agrupo las fallas de la ENCOLADORA
   RUNG wire#powerrail
      Contact( "Alarmas"."falla en rele de cadena" )
      wire#w1
      Coil( "Alarmas encoladora" )
   END_RUNG
   RUNG wire#powerrail
      Contact( "Alarmas"."Falla en sensor de encolado" )
   END_RUNG wire#w1
   RUNG wire#powerrail
      Contact( "Alarmas"."Sin pegamento en el depósito" )
   END_RUNG wire#w1
   // the same network as SCL:
   "Alarmas encoladora" := "Alarmas"."falla en rele de cadena" OR "Alarmas"."Falla en sensor de encolado" OR "Alarmas"."Sin pegamento en el depósito";
END_REGION

REGION Network 10: Serie de Alarmas
   RUNG wire#powerrail
      Contact( "Alarmas brazo de succión" )
      wire#w1
      Coil( "Serie de Alarmas" )
   END_RUNG
   RUNG wire#powerrail
      Contact( "Alarmas cinta" )
   END_RUNG wire#w1
   RUNG wire#powerrail
      Contact( "Alarmas emergencia y térmicas" )
   END_RUNG wire#w1
   RUNG wire#powerrail
      Contact( "Alarmas encoladora" )
   END_RUNG wire#w1
   RUNG wire#powerrail
      Contact( "Alarmas pusher" )
   END_RUNG wire#w1
   RUNG wire#powerrail
      Contact( "Alarmas salida y alim de cartones" )
   END_RUNG wire#w1
   RUNG wire#powerrail
      Contact( "Alarmas"."falla en rele de cadena" )
   END_RUNG wire#w1
   RUNG wire#powerrail
      Contact( "Alarmas"."caja cerrada en cadena" )
   END_RUNG wire#w1
   // the same network as SCL:
   "Serie de Alarmas" := "Alarmas brazo de succión" OR "Alarmas cinta" OR "Alarmas emergencia y térmicas" OR "Alarmas encoladora" OR "Alarmas pusher" OR "Alarmas salida y alim de cartones" OR "Alarmas"."falla en rele de cadena" OR "Alarmas"."caja cerrada en cadena";
END_REGION
END_FUNCTION

FUNCTION "Inversión de entradas" : Void   // FC5, LAD
TITLE = Invierte alguna entradas
{ S7_Optimized_Access := 'TRUE' }
VERSION : 0.1
BEGIN

REGION Network 1: Emergencia (Ventanas abiertas o Pulsador de emergencia)
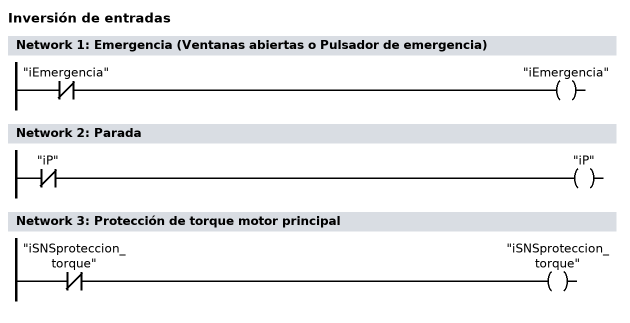
   RUNG wire#powerrail
      I_Contact( "iEmergencia" )
      Coil( "iEmergencia" )
   END_RUNG
   // the same network as SCL:
   "iEmergencia" := NOT "iEmergencia";
END_REGION

REGION Network 2: Parada
   RUNG wire#powerrail
      I_Contact( "iP" )
      Coil( "iP" )
   END_RUNG
   // the same network as SCL:
   "iP" := NOT "iP";
END_REGION

REGION Network 3: Protección de torque motor principal
   RUNG wire#powerrail
      I_Contact( "iSNSproteccion_torque" )
      Coil( "iSNSproteccion_torque" )
   END_RUNG
   // the same network as SCL:
   "iSNSproteccion_torque" := NOT "iSNSproteccion_torque";
END_REGION
END_FUNCTION

FUNCTION "Secuencia Principal" : Void   // FC6, LAD
TITLE = Secuencia Cinta Principal, Retenedores, Pinza, motor Pusher, cilindro Pusher
{ S7_Optimized_Access := 'TRUE' }
VERSION : 0.1
   VAR_TEMP   // added for the SCL form of the ladder/FBD networks
      _w1 : Bool;
   END_VAR
BEGIN

REGION Network 1: Muetra todos los estados para fines de diagnóstico.